// TIA Portal project "LabelProMax" (V16)

(* hardware
DEVICE "ET 200SP station_1"  ET 200SP-Station
   slot 0: "Rack_0"  Rack  6ES5 710-8MAx1
   slot 1: "PLC_label"  CPU 1512SP F-1 PN  6ES7 512-1SK01-0AB0  V2.8
      slot 32768: "PROFINET interface_1"  X1
         slot 32771: "Port_3"  X1 P3
   slot 2: "DI 8x24VDC HF_1"  DI 8x24VDC HF  6ES7 131-6BF00-0CA0  V1.2
      slot 1: "DI 8x24VDC HF_1"  DI 8x24VDC HF
   slot 3: "DI 8x24VDC HF_2"  DI 8x24VDC HF  6ES7 131-6BF00-0CA0  V1.2
      slot 1: "DI 8x24VDC HF_2"  DI 8x24VDC HF
   slot 4: "DQ 8x24VDC/0.5A HF_1"  DQ 8x24VDC/0.5A HF  6ES7 132-6BF00-0CA0  V1.2
      slot 1: "DQ 8x24VDC/0.5A HF_1"  DQ 8x24VDC/0.5A HF
   slot 5: "DQ 8x24VDC/0.5A HF_2"  DQ 8x24VDC/0.5A HF  6ES7 132-6BF00-0CA0  V1.2
      slot 1: "DQ 8x24VDC/0.5A HF_2"  DQ 8x24VDC/0.5A HF
   slot 6: "CM 4xIO-Link_1"  CM 4xIO-Link  6ES7 137-6BD00-0BA0  V2.1
      slot 1: "CM 4xIO-Link_1"  6ES7 137-6BD00-0BA0
   slot 7: "Server module_1"  Server module  6ES7 193-6PA00-0AA0  V1.0
      slot 1: "Server module_1"  Server module
   slot 127: "BA 2xRJ45"  BA 2xRJ45  6ES7 193-6AR00-0AA0  V0.0
      slot 32769: "Port_1"  X1 P1  6ES7 193-6AR00-0AA0
      slot 32770: "Port_2"  X1 P2  6ES7 193-6AR00-0AA0
DEVICE "HMI_label"  TP700 Comfort
   slot 0: "HMI_label"  TP700 Comfort  6AV2 124-0GC01-0AX0  16.0.0.0
   slot 1: "HMI_RT_1"  TP700 Comfort  6AV2 124-0GC01-0AX0  16.0.0.0
   slot 5: "HMI_label.IE_CP_1"  PROFINET Interface  16.0.0.0
      slot 1: "PROFINET Interface_1"  PROFINET Interface
         slot 1: "Port_1"  Port
         slot 2: "Port_2"  Port
   slot 7: "HMI_label.MPI/DP_CP_1"  MPI/DP Interface  16.0.0.0
*)

// ===== PLC "PLC_label"  CPU 1512SP F-1 PN =====

VAR_GLOBAL   // PLC tag table "Default tag table"
   "start" AT %I1.0 : Bool;   // 1=Start button pushed
   "stop" AT %I1.1 : Bool;   // 0=Stop button pushed (NC)
   "F1_F2" AT %I1.2 : Bool;   // 0=F1
   "reset" AT %I1.3 : Bool;   // 1=Reset button pushed
   "conv_centre" AT %I1.4 : Bool;   // 1=Carrier at conveyor centre
   "estop" AT %I1.5 : Bool;   // 0=Emergency stop button pushed (NC)
   "conv_start" AT %I1.6 : Bool;   // 1=Carrier at conveyor start
   "conv_end" AT %I1.7 : Bool;   // 1=Carrier at conveyor end
   "start_lamp" AT %Q1.0 : Bool;   // 1=Start lamp is lit
   "reset_lamp" AT %Q1.1 : Bool;   // 1=Reset lamp is lit
   "indicator_1" AT %Q1.2 : Bool;   // 1=Indicator Light 1 is lit
   "indicator_2" AT %Q1.3 : Bool;   // 1=Indicator Light 2 is lit
   "conv_fwd" AT %Q1.4 : Bool;   // 1=Move conveyor belt in clockwise rotation (to the right)
   "conv_bwd" AT %Q1.5 : Bool;   // 1=Move conveyor belt in counterclockwise rotation (to the left)
   "conv_inch" AT %Q1.6 : Bool;   // 1=Activate inch-travel of conveyor belt
   "stopper" AT %Q1.7 : Bool;   // 1=Move stopper cylinder to lower end position
END_VAR

VAR_GLOBAL   // PLC tag table "Tag table_1"
   "BG1" AT %I0.0 : Bool;
   "BG2" AT %I0.1 : Bool;
   "BG3" AT %I0.2 : Bool;
   "BG4" AT %I0.3 : Bool;
   "BG5" AT %I0.4 : Bool;
   "BG6" AT %I0.5 : Bool;
   "MB1" AT %Q0.0 : Bool;
   "MB3" AT %Q0.2 : Bool;
   "MB4" AT %Q0.3 : Bool;
   "MB5" AT %Q0.4 : Bool;
   "MB6" AT %Q0.5 : Bool;
   "MB7" AT %Q0.6 : Bool;
   "MA8" AT %Q0.7 : Bool;
END_VAR

DATA_BLOCK "base_Module_DB"   // DB1
{ S7_Optimized_Access := 'TRUE' }
VERSION : 0.1
// stored: InstanceOfName base_Module
"base_Module"
BEGIN
END_DATA_BLOCK

DATA_BLOCK "application_Module_DB"   // DB2
{ S7_Optimized_Access := 'TRUE' }
VERSION : 0.1
// stored: InstanceOfName application_Module
"application_Module"
BEGIN
END_DATA_BLOCK

DATA_BLOCK "Data_block_1"   // DB3
{ S7_Optimized_Access := 'TRUE' }
VERSION : 0.1
   VAR
      flag : Bool;
      state : Int;
      State1_Active : Bool;
      State2_Active : Bool;
      State3_Active : Bool;
      done : Bool;
      prev_done : Bool;
      "counter" : Int;
      run_timer : Real;
      prev_start : Bool;
      rfidDone : Bool;
      cycle_timer : TON_TIME;
      cycle_time_ms : DInt;
      total_runtime_ms : DInt;
      prev_rfidDone : Bool;
      timer_enable : Bool;
   END_VAR
BEGIN
END_DATA_BLOCK

DATA_BLOCK "LIOLink_RF200_ReadTag_DB"   // DB5
{ S7_Optimized_Access := 'FALSE' }
// stored: InstanceOfName LIOLink_RF200_ReadTag
"LIOLink_RF200_ReadTag"
BEGIN
END_DATA_BLOCK

DATA_BLOCK "RFID_Control"   // DB6
{ S7_Optimized_Access := 'TRUE' }
VERSION : 0.1
   VAR
      read : Bool := false;   // Execute a read of the RFID tag on rising edge
      write : Bool := false;
      length : Word := 16#1C;
      addrTag : Word := 16#00;
      hwID : Hw_SubModule := 261;
      portAddr : Int := 0;
      "version" : USInt := 11;
      readDone : Bool := false;
      writeDone : Bool := false;
      readPresence : Bool;
      writePresence : Bool;
   END_VAR
BEGIN
END_DATA_BLOCK

DATA_BLOCK "LIOLink_RF200_WriteTag_DB"   // DB7
{ S7_Optimized_Access := 'FALSE' }
// stored: InstanceOfName LIOLink_RF200_WriteTag
"LIOLink_RF200_WriteTag"
BEGIN
END_DATA_BLOCK

DATA_BLOCK "identData"   // DB8
{ S7_Optimized_Access := 'TRUE' }
VERSION : 0.1
   VAR
      readData : Array[0..31] of Byte;
      writeData : Array[0..31] of Byte;
   END_VAR
BEGIN
END_DATA_BLOCK

DATA_BLOCK "DB_MES_Comms"   // DB9
{ S7_Optimized_Access := 'TRUE' }
VERSION : 0.1
   VAR
      var1 : Bool;
      var2 : Int;
      var3 : Array[0..7] of Real;
      current_order_id : Int;
      station_state : Int;
      run_time : Real;
      total_count : Int;
      good_count : Int;
      completion_status : Bool;
      label_request : Bool;
      label_text : String[80];
      print_status : Bool;
      last_cycle_time : Real;
      cycle_done : Bool;
   END_VAR
BEGIN
END_DATA_BLOCK

DATA_BLOCK "state_Transition_Module_DB"   // DB10
{ S7_Optimized_Access := 'TRUE' }
VERSION : 0.1
// stored: InstanceOfName state_Transition_Module
"state_Transition_Module"
BEGIN
END_DATA_BLOCK

DATA_BLOCK "rfid_Current_Order_Module_DB"   // DB11
{ S7_Optimized_Access := 'TRUE' }
VERSION : 0.1
// stored: InstanceOfName rfid_Current_Order_Module
"rfid_Current_Order_Module"
BEGIN
END_DATA_BLOCK

FUNCTION_BLOCK "base_Module"   // FB1, GRAPH_PLUS
{ S7_Optimized_Access := 'TRUE' }
VERSION : 0.1
   VAR_INPUT
      OFF_SQ : Bool := false;   // Turn sequence off
      INIT_SQ : Bool := false;   // Set sequence to initial state
      ACK_EF : Bool := false;   // Acknowledge all errors and faults
      S_PREV : Bool := false;   // Output previous step in parameter S_NO
      S_NEXT : Bool := false;   // Indicate next step in parameter S_NO
      SW_AUTO : Bool := false;   // Automatic mode
      SW_TAP : Bool := false;   // Semiautomatic/switch with transition
      SW_TOP : Bool := false;   // Semiautomatic/ignore transition
      SW_MAN : Bool := false;   // Manual mode
      S_SEL : Int := 0;   // Select step to be output to S_NO
      S_ON : Bool := false;   // Activate step indicated in S_NO
      S_OFF : Bool := false;   // Deactivate step indicated S_NO
      T_PUSH : Bool := false;   // Enable transition to switch in semi automatic mode
   END_VAR
   VAR_OUTPUT
      S_NO : Int := 0;   // Step number
      S_MORE : Bool := false;   // More steps are available and can be shown in S_NO
      S_ACTIVE : Bool := false;   // Step indicated in S_NO is active
      ERR_FLT : Bool := false;   // Interlock or supervision group error
      AUTO_ON : Bool := false;   // Automatic mode is active
      TAP_ON : Bool := false;   // Semiautomatic mode/step with transition enabled
      TOP_ON : Bool := false;   // Semiautomatic mode/ignore transition enabled
      MAN_ON : Bool := false;   // Manual mode is active
   END_VAR
   VAR
      HMI_INFO : Array[0..8] of UInt;
      IF_PAR : G7_IfParPlus_V6;
      RT_DATA : G7_RTDataPlus_V6;   // Internal data area
      Trans1 : G7_TransitionPlus_V6;   // Transition structure
      Trans2 : G7_TransitionPlus_V6;   // Transition structure
      Trans3 : G7_TransitionPlus_V6;   // Transition structure
      Trans4 : G7_TransitionPlus_V6;   // Transition structure
      Trans5 : G7_TransitionPlus_V6;   // Transition structure
      Trans6 : G7_TransitionPlus_V6;   // Transition structure
      Trans7 : G7_TransitionPlus_V6;   // Transition structure
      Trans8 : G7_TransitionPlus_V6;   // Transition structure
      Trans9 : G7_TransitionPlus_V6;   // Transition structure
      Step1 : G7_StepPlus_V6;   // Step structure
      Step2 : G7_StepPlus_V6;   // Step structure
      Step3 : G7_StepPlus_V6;   // Step structure
      Step4 : G7_StepPlus_V6;   // Step structure
      Step5 : G7_StepPlus_V6;   // Step structure
      Step6 : G7_StepPlus_V6;   // Step structure
      Step7 : G7_StepPlus_V6;   // Step structure
      Step8 : G7_StepPlus_V6;   // Step structure
      Step9 : G7_StepPlus_V6;   // Step structure
      SINI : Array[0..1] of USInt;
      LSTT : Array[0..8] of USInt;
      ATAJ : Array[0..8] of USInt;
      ATAB : Array[0..8] of USInt;
      PSTT : Array[0..8] of USInt;
      NSTT : Array[0..8] of USInt;
      ASSJ : Array[0..8] of USInt;
      ASSB : Array[0..8] of USInt;
      PTTS : Array[0..8] of USInt;
      NTTS : Array[0..8] of USInt;
      SW_SQTS : Array[0..8] of USInt;
      SWITCH : Array[0..0] of USInt;
      TVX : Array[0..1] of USInt;
      TTX : Array[0..1] of USInt;
      TSX : Array[0..1] of USInt;
      S00X : Array[0..1] of USInt;
      SOFFX : Array[0..1] of USInt;
      SONX : Array[0..1] of USInt;
      SAX : Array[0..1] of USInt;
      SERRX : Array[0..9] of USInt;
      SMX : Array[0..9] of USInt;
      S0X : Array[0..9] of USInt;
      S1X : Array[0..9] of USInt;
      IL_ALARM_INST : Diag_Alarm;
      SUP_ALARM_INST : Diag_Alarm;
      STEP_TIME_ALARM_INST : Diag_Alarm;
      IEC_TIMER_INST : IEC_TIMER;
      TRANSACTION_FLAG : Bool := false;
   END_VAR
   // SINI[0] := 2;
   // LSTT[0] := 255;
   // LSTT[1] := 255;
   // LSTT[2] := 255;
   // ATAJ[1] := 1;
   // ATAJ[2] := 2;
   // ATAJ[3] := 3;
   // ATAB[1] := 1;
   // ATAB[2] := 2;
   // ATAB[3] := 3;
   // PSTT[1] := 1;
   // PSTT[2] := 2;
   // PSTT[3] := 5;
   // NSTT[0] := 1;
   // NSTT[1] := 6;
   // NSTT[2] := 3;
   // ASSJ[1] := 1;
   // ASSJ[2] := 2;
   // ASSJ[3] := 3;
   // ASSB[1] := 1;
   // ASSB[2] := 2;
   // ASSB[3] := 3;
   // PTTS[0] := 255;
   // PTTS[2] := 8;
   // PTTS[3] := 2;
   // NTTS[1] := 1;
   // NTTS[2] := 2;
   // NTTS[3] := 5;
   // TVX[0] := 16#1;
   // TTX[0] := 16#1;
   // TSX[0] := 16#1;
   // S00X[0] := 16#1;
   // SOFFX[0] := 16#1;
   // SONX[0] := 16#1;
   // SAX[0] := 16#1;
   // SERRX[0] := 16#1;
   // SMX[0] := 16#1;
   // S0X[0] := 16#1;
   // S1X[0] := 16#1;
   // LSTT[3] := 255;
   // ATAJ[4] := 4;
   // ATAB[4] := 4;
   // PSTT[4] := 4;
   // NSTT[3] := 4;
   // ASSJ[4] := 4;
   // ASSB[4] := 4;
   // PTTS[4] := 3;
   // NTTS[4] := 4;
   // LSTT[5] := 255;
   // ATAJ[5] := 5;
   // ATAB[5] := 5;
   // PSTT[5] := 3;
   // NSTT[5] := 5;
   // ASSJ[5] := 5;
   // ASSB[5] := 5;
   // PTTS[5] := 5;
   // NTTS[5] := 3;
   // LSTT[6] := 255;
   // ATAJ[6] := 6;
   // ATAB[6] := 6;
   // PSTT[6] := 6;
   // NSTT[6] := 7;
   // ASSJ[6] := 6;
   // ASSB[6] := 6;
   // PTTS[6] := 1;
   // NTTS[6] := 6;
   // LSTT[7] := 255;
   // LSTT[8] := 255;
   // ATAJ[7] := 7;
   // ATAJ[8] := 8;
   // ATAB[7] := 7;
   // ATAB[8] := 8;
   // PSTT[7] := 7;
   // PSTT[8] := 8;
   // NSTT[7] := 8;
   // NSTT[8] := 2;
   // ASSJ[7] := 7;
   // ASSJ[8] := 8;
   // ASSB[7] := 7;
   // ASSB[8] := 8;
   // PTTS[7] := 6;
   // PTTS[8] := 7;
   // NTTS[7] := 7;
   // NTTS[8] := 8;
BEGIN
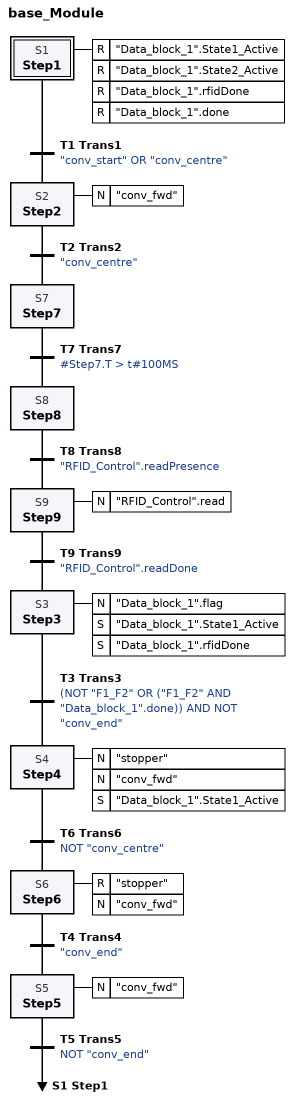
   // sequencer 1
   INITIAL_STEP Step1:   // S1, max time T#10S, warning time T#7S
              R    "Data_block_1".State1_Active
              R    "Data_block_1".State2_Active
              R    "Data_block_1".rfidDone
              R    "Data_block_1".done
   END_STEP
   TRANSITION Trans1 FROM Step1 TO Step2   // T1
      := "conv_start" OR "conv_centre";
   END_TRANSITION
   STEP Step2:   // S2, max time T#10S, warning time T#7S
              N    "conv_fwd"
   END_STEP
   TRANSITION Trans2 FROM Step2 TO Step7   // T2
      := "conv_centre";
   END_TRANSITION
   STEP Step3:   // S3, max time T#10S, warning time T#7S
              N    "Data_block_1".flag
              S    "Data_block_1".State1_Active
              S    "Data_block_1".rfidDone
   END_STEP
   TRANSITION Trans3 FROM Step3 TO Step4   // T3
      := (NOT "F1_F2" OR ("F1_F2" AND "Data_block_1".done)) AND NOT "conv_end";
   END_TRANSITION
   STEP Step4:   // S4, max time T#10S, warning time T#7S
              N    "stopper"
              N    "conv_fwd"
              S    "Data_block_1".State1_Active
   END_STEP
   TRANSITION Trans6 FROM Step4 TO Step6   // T6
      := NOT "conv_centre";
   END_TRANSITION
   STEP Step5:   // S5, max time T#10S, warning time T#7S
              N    "conv_fwd"
   END_STEP
   TRANSITION Trans5 FROM Step5 TO Step1   // T5, jump
      := NOT "conv_end";
   END_TRANSITION
   STEP Step6:   // S6, max time T#10S, warning time T#7S
              R    "stopper"
              N    "conv_fwd"
   END_STEP
   TRANSITION Trans4 FROM Step6 TO Step5   // T4
      := "conv_end";
   END_TRANSITION
   STEP Step7:   // S7, max time T#10S, warning time T#7S
   END_STEP
   TRANSITION Trans7 FROM Step7 TO Step8   // T7
      := #Step7.T > t#100MS;
   END_TRANSITION
   STEP Step8:   // S8, max time T#10S, warning time T#7S
   END_STEP
   TRANSITION Trans8 FROM Step8 TO Step9   // T8
      := "RFID_Control".readPresence;
   END_TRANSITION
   STEP Step9:   // S9, max time T#10S, warning time T#7S
              N    "RFID_Control".read
   END_STEP
   TRANSITION Trans9 FROM Step9 TO Step3   // T9
      := "RFID_Control".readDone;
   END_TRANSITION
END_FUNCTION_BLOCK

FUNCTION_BLOCK "application_Module"   // FB2, GRAPH_PLUS
{ S7_Optimized_Access := 'TRUE' }
VERSION : 0.1
   VAR_INPUT
      OFF_SQ : Bool := false;   // Turn sequence off
      INIT_SQ : Bool := false;   // Set sequence to initial state
      ACK_EF : Bool := false;   // Acknowledge all errors and faults
      S_PREV : Bool := false;   // Output previous step in parameter S_NO
      S_NEXT : Bool := false;   // Indicate next step in parameter S_NO
      SW_AUTO : Bool := false;   // Automatic mode
      SW_TAP : Bool := false;   // Semiautomatic/switch with transition
      SW_TOP : Bool := false;   // Semiautomatic/ignore transition
      SW_MAN : Bool := false;   // Manual mode
      S_SEL : Int := 0;   // Select step to be output to S_NO
      S_ON : Bool := false;   // Activate step indicated in S_NO
      S_OFF : Bool := false;   // Deactivate step indicated S_NO
      T_PUSH : Bool := false;   // Enable transition to switch in semi automatic mode
   END_VAR
   VAR_OUTPUT
      S_NO : Int := 0;   // Step number
      S_MORE : Bool := false;   // More steps are available and can be shown in S_NO
      S_ACTIVE : Bool := false;   // Step indicated in S_NO is active
      ERR_FLT : Bool := false;   // Interlock or supervision group error
      AUTO_ON : Bool := false;   // Automatic mode is active
      TAP_ON : Bool := false;   // Semiautomatic mode/step with transition enabled
      TOP_ON : Bool := false;   // Semiautomatic mode/ignore transition enabled
      MAN_ON : Bool := false;   // Manual mode is active
   END_VAR
   VAR
      HMI_INFO : Array[0..8] of UInt;
      IF_PAR : G7_IfParPlus_V6;
      RT_DATA : G7_RTDataPlus_V6;   // Internal data area
      Trans1 : G7_TransitionPlus_V6;   // Transition structure
      Trans2 : G7_TransitionPlus_V6;   // Transition structure
      Trans3 : G7_TransitionPlus_V6;   // Transition structure
      Trans4 : G7_TransitionPlus_V6;   // Transition structure
      Trans5 : G7_TransitionPlus_V6;   // Transition structure
      Trans6 : G7_TransitionPlus_V6;   // Transition structure
      Trans7 : G7_TransitionPlus_V6;   // Transition structure
      Trans8 : G7_TransitionPlus_V6;   // Transition structure
      Trans9 : G7_TransitionPlus_V6;   // Transition structure
      Trans10 : G7_TransitionPlus_V6;   // Transition structure
      Trans11 : G7_TransitionPlus_V6;   // Transition structure
      Step1 : G7_StepPlus_V6;   // Step structure
      Step2 : G7_StepPlus_V6;   // Step structure
      Step3 : G7_StepPlus_V6;   // Step structure
      Step4 : G7_StepPlus_V6;   // Step structure
      Step5 : G7_StepPlus_V6;   // Step structure
      Step6 : G7_StepPlus_V6;   // Step structure
      Step7 : G7_StepPlus_V6;   // Step structure
      Step8 : G7_StepPlus_V6;   // Step structure
      Step9 : G7_StepPlus_V6;   // Step structure
      Step10 : G7_StepPlus_V6;   // Step structure
      Step11 : G7_StepPlus_V6;   // Step structure
      SINI : Array[0..1] of USInt;
      LSTT : Array[0..10] of USInt;
      ATAJ : Array[0..10] of USInt;
      ATAB : Array[0..10] of USInt;
      PSTT : Array[0..10] of USInt;
      NSTT : Array[0..10] of USInt;
      ASSJ : Array[0..10] of USInt;
      ASSB : Array[0..10] of USInt;
      PTTS : Array[0..10] of USInt;
      NTTS : Array[0..10] of USInt;
      SW_SQTS : Array[0..10] of USInt;
      SWITCH : Array[0..0] of USInt;
      TVX : Array[0..1] of USInt;
      TTX : Array[0..1] of USInt;
      TSX : Array[0..1] of USInt;
      S00X : Array[0..1] of USInt;
      SOFFX : Array[0..1] of USInt;
      SONX : Array[0..1] of USInt;
      SAX : Array[0..1] of USInt;
      SERRX : Array[0..11] of USInt;
      SMX : Array[0..11] of USInt;
      S0X : Array[0..11] of USInt;
      S1X : Array[0..11] of USInt;
      IL_ALARM_INST : Diag_Alarm;
      SUP_ALARM_INST : Diag_Alarm;
      STEP_TIME_ALARM_INST : Diag_Alarm;
      IEC_TIMER_INST : IEC_TIMER;
      TRANSACTION_FLAG : Bool := false;
   END_VAR
   // SINI[0] := 2;
   // LSTT[0] := 255;
   // LSTT[1] := 255;
   // LSTT[2] := 255;
   // LSTT[3] := 255;
   // LSTT[4] := 255;
   // LSTT[5] := 255;
   // LSTT[6] := 255;
   // LSTT[7] := 255;
   // LSTT[8] := 255;
   // LSTT[9] := 255;
   // ATAJ[1] := 1;
   // ATAJ[2] := 2;
   // ATAJ[3] := 3;
   // ATAJ[4] := 4;
   // ATAJ[5] := 5;
   // ATAJ[6] := 6;
   // ATAJ[7] := 7;
   // ATAJ[8] := 8;
   // ATAJ[9] := 9;
   // ATAJ[10] := 10;
   // ATAB[1] := 1;
   // ATAB[2] := 2;
   // ATAB[3] := 3;
   // ATAB[4] := 4;
   // ATAB[5] := 5;
   // ATAB[6] := 6;
   // ATAB[7] := 7;
   // ATAB[8] := 8;
   // ATAB[9] := 9;
   // ATAB[10] := 10;
   // PSTT[1] := 1;
   // PSTT[2] := 2;
   // PSTT[3] := 3;
   // PSTT[4] := 4;
   // PSTT[5] := 5;
   // PSTT[6] := 6;
   // PSTT[7] := 7;
   // PSTT[8] := 8;
   // PSTT[9] := 9;
   // PSTT[10] := 10;
   // NSTT[0] := 1;
   // NSTT[1] := 2;
   // NSTT[2] := 3;
   // NSTT[3] := 4;
   // NSTT[4] := 5;
   // NSTT[5] := 6;
   // NSTT[6] := 7;
   // NSTT[7] := 8;
   // NSTT[8] := 9;
   // NSTT[9] := 10;
   // ASSJ[1] := 1;
   // ASSJ[2] := 2;
   // ASSJ[3] := 3;
   // ASSJ[4] := 4;
   // ASSJ[5] := 5;
   // ASSJ[6] := 6;
   // ASSJ[7] := 7;
   // ASSJ[8] := 8;
   // ASSJ[9] := 9;
   // ASSJ[10] := 10;
   // ASSB[1] := 1;
   // ASSB[2] := 2;
   // ASSB[3] := 3;
   // ASSB[4] := 4;
   // ASSB[5] := 5;
   // ASSB[6] := 6;
   // ASSB[7] := 7;
   // ASSB[8] := 8;
   // ASSB[9] := 9;
   // ASSB[10] := 10;
   // PTTS[0] := 255;
   // PTTS[2] := 1;
   // PTTS[3] := 2;
   // PTTS[4] := 3;
   // PTTS[5] := 4;
   // PTTS[6] := 5;
   // PTTS[7] := 6;
   // PTTS[8] := 7;
   // PTTS[9] := 8;
   // PTTS[10] := 9;
   // NTTS[1] := 1;
   // NTTS[2] := 2;
   // NTTS[3] := 3;
   // NTTS[4] := 4;
   // NTTS[5] := 5;
   // NTTS[6] := 6;
   // NTTS[7] := 7;
   // NTTS[8] := 8;
   // NTTS[9] := 9;
   // NTTS[10] := 10;
   // TVX[0] := 16#1;
   // TTX[0] := 16#1;
   // TSX[0] := 16#1;
   // S00X[0] := 16#1;
   // SOFFX[0] := 16#1;
   // SONX[0] := 16#1;
   // SAX[0] := 16#1;
   // SERRX[0] := 16#1;
   // SMX[0] := 16#1;
   // S0X[0] := 16#1;
   // S1X[0] := 16#1;
BEGIN
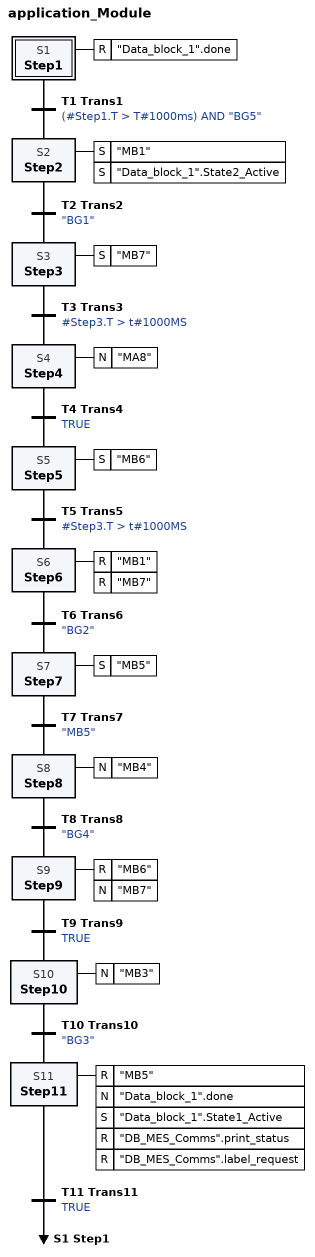
   // sequencer 1
   INITIAL_STEP Step1:   // S1, max time T#10S, warning time T#7S
              R    "Data_block_1".done
   END_STEP
   TRANSITION Trans1 FROM Step1 TO Step2   // T1
      := (#Step1.T > T#1000ms) AND "BG5";
   END_TRANSITION
   STEP Step2:   // S2, max time T#10S, warning time T#7S
              S    "MB1"
              S    "Data_block_1".State2_Active
   END_STEP
   TRANSITION Trans2 FROM Step2 TO Step3   // T2
      := "BG1";
   END_TRANSITION
   STEP Step3:   // S3, max time T#10S, warning time T#7S
              S    "MB7"
   END_STEP
   TRANSITION Trans3 FROM Step3 TO Step4   // T3
      := #Step3.T > t#1000MS;
   END_TRANSITION
   STEP Step4:   // S4, max time T#10S, warning time T#7S
              N    "MA8"
   END_STEP
   TRANSITION Trans4 FROM Step4 TO Step5   // T4
      := TRUE;
   END_TRANSITION
   STEP Step5:   // S5, max time T#10S, warning time T#7S
              S    "MB6"
   END_STEP
   TRANSITION Trans5 FROM Step5 TO Step6   // T5
      := #Step3.T > t#1000MS;
   END_TRANSITION
   STEP Step6:   // S6, max time T#10S, warning time T#7S
              R    "MB1"
              R    "MB7"
   END_STEP
   TRANSITION Trans6 FROM Step6 TO Step7   // T6
      := "BG2";
   END_TRANSITION
   STEP Step7:   // S7, max time T#10S, warning time T#7S
              S    "MB5"
   END_STEP
   TRANSITION Trans7 FROM Step7 TO Step8   // T7
      := "MB5";
   END_TRANSITION
   STEP Step8:   // S8, max time T#10S, warning time T#7S
              N    "MB4"
   END_STEP
   TRANSITION Trans8 FROM Step8 TO Step9   // T8
      := "BG4";
   END_TRANSITION
   STEP Step9:   // S9, max time T#10S, warning time T#7S
              R    "MB6"
              N    "MB7"
   END_STEP
   TRANSITION Trans9 FROM Step9 TO Step10   // T9
      := TRUE;
   END_TRANSITION
   STEP Step10:   // S10, max time T#10S, warning time T#7S
              N    "MB3"
   END_STEP
   TRANSITION Trans10 FROM Step10 TO Step11   // T10
      := "BG3";
   END_TRANSITION
   STEP Step11:   // S11, max time T#10S, warning time T#7S
              R    "MB5"
              N    "Data_block_1".done
              S    "Data_block_1".State1_Active
              R    "DB_MES_Comms".print_status
              R    "DB_MES_Comms".label_request
   END_STEP
   TRANSITION Trans11 FROM Step11 TO Step1   // T11, jump
      := TRUE;
   END_TRANSITION
END_FUNCTION_BLOCK

FUNCTION_BLOCK "state_Transition_Module"   // FB4, SCL
{ S7_Optimized_Access := 'TRUE' }
VERSION : 0.1
BEGIN
   IF "Data_block_1".State2_Active THEN
       "Data_block_1".state := 2;
       "DB_MES_Comms".station_state := "Data_block_1".state;
   ELSIF "Data_block_1".State1_Active THEN
       "Data_block_1".state := 1;
       "DB_MES_Comms".station_state := "Data_block_1".state;
   ELSE
       "Data_block_1".state := 0;
       "DB_MES_Comms".station_state := "Data_block_1".state;
   END_IF;
END_FUNCTION_BLOCK

ORGANIZATION_BLOCK "Main"   // OB1, LAD, ProgramCycle
TITLE = "Main Program Sweep (Cycle)"
{ S7_Optimized_Access := 'TRUE' }
VERSION : 0.1
   VAR_INPUT
      Initial_Call : Bool;   // Initial call of this OB
      Remanence : Bool;   // =True, if remanent data are available
   END_VAR
   VAR_TEMP
      run_time_ms : Real;
   END_VAR
BEGIN

REGION Network 1: Execution of Converyor belt start stop logic in Block_1 [FB1]
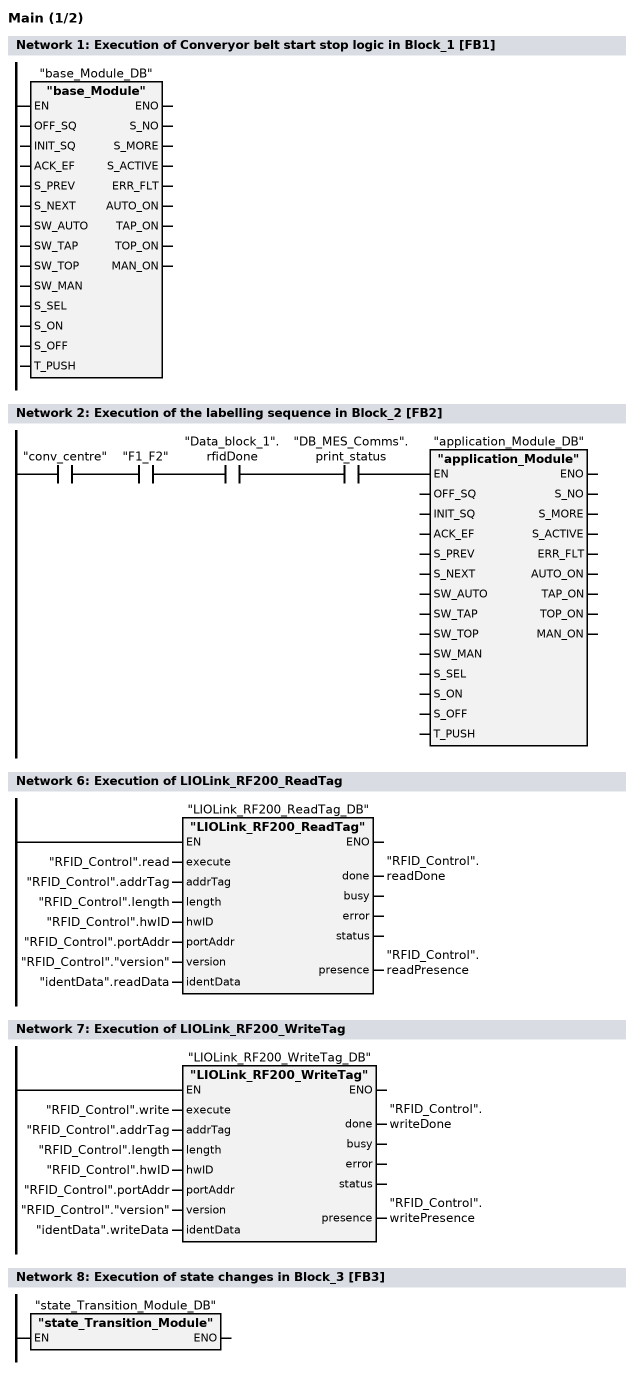
   RUNG wire#powerrail
      "base_Module_DB"(OFF_SQ :=, INIT_SQ :=, ACK_EF :=, S_PREV :=, S_NEXT :=, SW_AUTO :=, SW_TAP :=, SW_TOP :=, SW_MAN :=, S_SEL :=, S_ON :=, S_OFF :=, T_PUSH :=, S_NO =>, S_MORE =>, S_ACTIVE =>, ERR_FLT =>, AUTO_ON =>, TAP_ON =>, TOP_ON =>, MAN_ON =>)
   END_RUNG
   // the same network as SCL:
   "base_Module_DB"();   // "base_Module"
END_REGION

REGION Network 2: Execution of the labelling sequence in Block_2 [FB2]
   RUNG wire#powerrail
      Contact( "conv_centre" )
      Contact( "F1_F2" )
      Contact( "Data_block_1".rfidDone )
      Contact( "DB_MES_Comms".print_status )
      "application_Module_DB"(OFF_SQ :=, INIT_SQ :=, ACK_EF :=, S_PREV :=, S_NEXT :=, SW_AUTO :=, SW_TAP :=, SW_TOP :=, SW_MAN :=, S_SEL :=, S_ON :=, S_OFF :=, T_PUSH :=, S_NO =>, S_MORE =>, S_ACTIVE =>, ERR_FLT =>, AUTO_ON =>, TAP_ON =>, TOP_ON =>, MAN_ON =>)
   END_RUNG
   // the same network as SCL:
   IF "conv_centre" AND "F1_F2" AND "Data_block_1".rfidDone AND "DB_MES_Comms".print_status THEN
       "application_Module_DB"();   // "application_Module"
   END_IF;
END_REGION

REGION Network 3 (SCL): Total Count
   IF "Data_block_1".State1_Active AND NOT "Data_block_1".prev_start AND "F1_F2" = TRUE THEN

       "DB_MES_Comms".total_count := "DB_MES_Comms".total_count + 1;

   END_IF;

   "Data_block_1".prev_start := "Data_block_1".State1_Active;
END_REGION

REGION Network 4 (SCL): Good Count
   IF "Data_block_1".done AND NOT "Data_block_1".prev_done AND "F1_F2" = TRUE THEN

       "DB_MES_Comms".good_count := "DB_MES_Comms".good_count + 1;

   END_IF;

   "Data_block_1".prev_done := "Data_block_1".done;
END_REGION

REGION Network 5 (SCL): Completion Status of the orders sent by MES (not in reality\)
   IF "DB_MES_Comms".total_count >= 10 THEN
       "DB_MES_Comms".completion_status := TRUE;
   ELSE
       "DB_MES_Comms".completion_status := FALSE;
   END_IF;
END_REGION

REGION Network 6: Execution of LIOLink_RF200_ReadTag
   RUNG wire#powerrail
      "LIOLink_RF200_ReadTag_DB"(execute := "RFID_Control".read, addrTag := "RFID_Control".addrTag, length := "RFID_Control".length, hwID := "RFID_Control".hwID, portAddr := "RFID_Control".portAddr, "version" := "RFID_Control"."version", identData := "identData".readData, done => "RFID_Control".readDone, busy =>, error =>, status =>, presence => "RFID_Control".readPresence)
   END_RUNG
   // the same network as SCL:
   "LIOLink_RF200_ReadTag_DB"(execute := "RFID_Control".read,   // "LIOLink_RF200_ReadTag"
                           addrTag := "RFID_Control".addrTag,
                           length := "RFID_Control".length,
                           hwID := "RFID_Control".hwID,
                           portAddr := "RFID_Control".portAddr,
                           "version" := "RFID_Control"."version",
                           identData := "identData".readData,
                           done => "RFID_Control".readDone,
                           presence => "RFID_Control".readPresence);
END_REGION

REGION Network 7: Execution of LIOLink_RF200_WriteTag
   RUNG wire#powerrail
      "LIOLink_RF200_WriteTag_DB"(execute := "RFID_Control".write, addrTag := "RFID_Control".addrTag, length := "RFID_Control".length, hwID := "RFID_Control".hwID, portAddr := "RFID_Control".portAddr, "version" := "RFID_Control"."version", identData := "identData".writeData, done => "RFID_Control".writeDone, busy =>, error =>, status =>, presence => "RFID_Control".writePresence)
   END_RUNG
   // the same network as SCL:
   "LIOLink_RF200_WriteTag_DB"(execute := "RFID_Control".write,   // "LIOLink_RF200_WriteTag"
                           addrTag := "RFID_Control".addrTag,
                           length := "RFID_Control".length,
                           hwID := "RFID_Control".hwID,
                           portAddr := "RFID_Control".portAddr,
                           "version" := "RFID_Control"."version",
                           identData := "identData".writeData,
                           done => "RFID_Control".writeDone,
                           presence => "RFID_Control".writePresence);
END_REGION

REGION Network 8: Execution of state changes in Block_3 [FB3]
   RUNG wire#powerrail
      "state_Transition_Module_DB"()
   END_RUNG
   // the same network as SCL:
   "state_Transition_Module_DB"();   // "state_Transition_Module"
END_REGION

REGION Network 9 (SCL): Start Timer on RFID Done
   IF "Data_block_1".rfidDone AND NOT "Data_block_1".prev_rfidDone THEN
       "Data_block_1".timer_enable := TRUE;
   END_IF;

   "Data_block_1".prev_rfidDone := "Data_block_1".rfidDone;
END_REGION

REGION Network 10 (SCL): Cycle Timer (Controlled)
   "Data_block_1".cycle_timer(
                              IN := "Data_block_1".timer_enable,
                              PT := T#9999s
   );
END_REGION

REGION Network 11 (SCL): Stop Timer + Accumulate Runtime
   IF "Data_block_1".done AND NOT "Data_block_1".prev_done THEN

       "Data_block_1".timer_enable := false;

       "Data_block_1".cycle_time_ms := "Data_block_1".cycle_timer.ET;

       "Data_block_1".total_runtime_ms := "Data_block_1".total_runtime_ms + "Data_block_1".cycle_time_ms;

       "DB_MES_Comms".last_cycle_time := DINT_TO_REAL("Data_block_1".cycle_time_ms) / 1000.0;

       "DB_MES_Comms".cycle_done := TRUE;

   END_IF;

   "Data_block_1".prev_done := "Data_block_1".done;
END_REGION

REGION Network 12 (SCL): Reset cycle_done Signal
   IF "DB_MES_Comms".cycle_done THEN
       "DB_MES_Comms".cycle_done := FALSE;
   END_IF;
END_REGION

REGION Network 13 (SCL): MES Publish
   "DB_MES_Comms".run_time := DINT_TO_REAL("Data_block_1".total_runtime_ms) / 1000.0;
   "DB_MES_Comms".station_state := "Data_block_1".state;
END_REGION

REGION Network 14: Activate DB_MES_Comms.label_request when LIO...ReadTag_DB.done is true and DB...ms.print_status is false
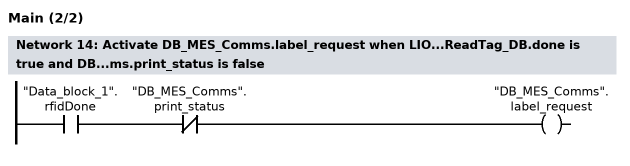
   RUNG wire#powerrail
      Contact( "Data_block_1".rfidDone )
      I_Contact( "DB_MES_Comms".print_status )
      Coil( "DB_MES_Comms".label_request )
   END_RUNG
   // the same network as SCL:
   "DB_MES_Comms".label_request := "Data_block_1".rfidDone AND NOT "DB_MES_Comms".print_status;
END_REGION
END_ORGANIZATION_BLOCK

// folder: LIOLink/S7-1200/1500/Device-specific blocks/SIMATIC RF200

FUNCTION_BLOCK "LIOLink_RF200_ReadTag"   // FB3, SCL
TITLE = LIOLink_RF200_ReadTag
{ S7_Optimized_Access := 'FALSE' }
// Reads tags from SIMATIC RF200 readers via IO-Link
   VAR_INPUT
      execute : Bool;   // Execute function
      addrTag : Word;   // Start address of data on tag
      length : Word;   // Length of data to be read
      hwID : Hw_SubModule;   // Hardware identifier of IO-Link communication module
      portAddr : Int;   // Start address of port
      "version" : USInt := 11;   // IO-Link version of the reader; 11: IO-Link V1.1, 10: IO-Link V1.0
   END_VAR
   VAR_OUTPUT
      done : Bool;
      busy : Bool;
      error : Bool;
      status : DWord;
      statusWord AT status : Array[0..1] of Word;
      presence : Bool;
   END_VAR
   VAR_IN_OUT
      identData : Variant;
   END_VAR
   VAR
      statPae : Array[0..27] of Byte;
      statStatusByte : Byte;
      statStatusBit AT statStatusByte : Array[0..7] of Bool;
      statPresence : Bool;
      statState : Int;
      statIdleState : Int;
      statTelegramState : Int := 1;
      statReadState : Int := 2;
      statErrorState : Int := 3;
      statAddr : Word;
      statAddrRead AT statAddr : Array[0..1] of Byte;
      statOffset : Int;
      statExecuteReq : Bool;
      statLength : DInt;
      statDat : Array[0..31] of Byte;
      statRecDat : Array[0..31] of Byte;
      statAddrOffset : Int;
      statPresenceFF : Bool;
      InstTonrTime : TONR_TIME;
      statTimerIn : Bool;
      statTimerR : Bool;
      statTimerPt : Time := t#5s;
      statReadData : Array[0..1999] of Byte;
      statCountCopyPae : DInt;
      statBusy : Bool;
      statDone : Bool;
      statReturnMoveBlkVar : Int;
      statDiffToIOsizeNetto : Int;
      InstSetIoPart : SETIO_PART;
      statIoPartError : Bool;
      statIoPartStatus : DWord;
      InstGetIoPart : GETIO_PART;
      statIOsize : USInt;
      statIOsizeNetto : USInt;
   END_VAR
   VAR_TEMP
      tempError : Bool;
      tempStatus : DWord;
      tempStatus_W AT tempStatus : Array[0..1] of Word;
   END_VAR
   VAR CONSTANT
      IOL_V10 : USInt := 10;   // Identifier IO-Link version 1.0
      IOL_V11 : USInt := 11;   // Identifier IO-Link version 1.1
      LEN_DATA_V10 : USInt := 8;   // Length of user data for IO-Link version 1.0
      LEN_DATA_V11 : USInt := 32;   // Length of user data for IO-Link version 1.1
   END_VAR
BEGIN
   REGION BLOCK INFO HEADER
     //===============================================================================
     // Siemens / (c)Copyright 2020
     //-------------------------------------------------------------------------------
     // Title:            LIOLink_RF200_ReadTag
     // Function:         Reads tags from SIMATIC RF200 readers via IO-Link
     // Library:          LIOLink
     // Author:           Siemens Industry Online Support
     // Tested with:      CPU 1513-1 PN FW 2.8
     // Engineering:      TIA Portal V16
     // Restrictions:     --
     // Requirements:     --
     //-------------------------------------------------------------------------------
     // Change log table:
     // Version  | Date       | Expert in charge       | Changes applied
     //----------|------------|------------------------|------------------------------
     // 01.00.00 | 01.07.2013 | Online Support         | First release
     // 01.01.00 | 01.12.2016 | Online Support         | Upgraded to TIA Portal V14
     // 02.00.00 | 01.09.2017 | Online Support         | Upgraded to TIA Portal V14 SP1
     //                                                | Implemented Programming styleguide
     //                                                | Added support for IO-Link V1.1 readers
     // 02.01.00 | 01.12.2017 | Online Support         | Bug fixes and performance improvements
     // 02.02.00 | 01.03.2020 | Online Support         | Upgraded to TIA Portal V16
     // 02.03.00 | 22.09.2020 | Online Support         | Integrated FB into LIOLink library
     //                                                | Renamed FB to LIOLink_RF200_ReadTag
     //                                                | Combined FBs for IO-Link V1.0 and V1.1
     //                                                | Minor bug fixes
     //===============================================================================
   END_REGION

   IF #version = #IOL_V11 THEN                               //determine IO-Link reader version (1.0/1.1) to set offsets
       #statIOsize := #LEN_DATA_V11;
       #statIOsizeNetto := #LEN_DATA_V11 - 4;
   ELSE
       #statIOsize := #LEN_DATA_V10;
       #statIOsizeNetto := #LEN_DATA_V10 - 4;
   END_IF;

   #statAddrOffset := #portAddr;                           //start adress of port
   #InstGetIoPart(ID     := #hwID,
                  OFFSET := #statAddrOffset,
                  LEN    := #statIOsize,
                  STATUS => #statIoPartStatus,
                  ERROR  => #statIoPartError,
                  INPUTS := #statRecDat);

   #statStatusByte := #statRecDat[0];         //Status Byte
   #statPresence := #statStatusBit[5];                     //Presence bit. Transponder on field
   #presence := #statPresence;

   IF NOT #execute THEN
       #statDone := false;
       #statBusy := false;
       #done := false;
       #busy := false;
       #error := false;
       #status := 0;
   ELSE
       #done := #statDone;
       #busy := #statBusy;
   END_IF;

   IF #execute AND #execute <> #statExecuteReq THEN        //Positive edge for d#reading of data
       IF NOT #statBusy THEN
           #statAddr := #addrTag;                                    //Transpoder Address
           #statDiffToIOsizeNetto := WORD_TO_INT(#length) MOD #statIOsizeNetto;
           #statLength := #length;                                 //Length of read Dat
           #statBusy := TRUE;
           #statDone := FALSE;                                     //reset all the output parameters                                   
           #error := FALSE;
           #status := 0;
           #statOffset := 0;                                       //offset of puffer must be reseted
           #statState := #statReadState;                           //next step >> send read command
           #statCountCopyPae := 0;
           FILL_BLK(IN    := 0,                                    //Reset read buffer
                    COUNT := CountOfElements(#identData),
                    OUT   => #statReadData[0]);
       ELSE
           #tempStatus_W[1] := 16#8102;                            //block is still active
           #tempStatus_W[0] := 16#0001;                            //Error identifier for block errors
           #status := #tempStatus;
           #statState := #statErrorState;
       END_IF;
       IF #length < 0 THEN
           #tempStatus_W[1] := 16#8104;                             //length too short
           #tempStatus_W[0] := 16#0001;                             //identifier rfid errors
           #status := #tempStatus;
           #statState := #statErrorState;
       END_IF;
   END_IF;
   #statExecuteReq := #execute;

   IF NOT #presence AND #presence <> #statPresenceFF THEN   //the tag has left the antenna  field
       IF NOT #statDone THEN
           #statTimerIn := true;                              //wait 5 sec
           #statTimerR := false;
       END_IF;
   END_IF;
   #statPresenceFF := #presence;
   IF #presence THEN
       #statTimerR := true;
       #statTimerIn := false;
   END_IF;
   //-----------------------------------------------------------------------------------------------------//
   //------------------------------------------start of state machine------------------------------------//
   //-----------------------------------------------------------------------------------------------------//
   CASE #statState OF
       0://IDLE
           #statBusy := false;
           #statTimerIn := false;

           (*
           // #statAdr := 0;
           // #statDat[0] := 16#0;                      //Set read command
           // #statDat[2] := #statAdrRead[0];             //Adr-H
           // #statDat[3] := #statAdrRead[1];             //Adr-L
           // #InstSetIoPart(ID:=#hwId,
           //                OFFSET:=#statAdrOffset,
           //                LEN:=8,
           //                STATUS=>#statIoPartStatus,
           //                ERROR=>#statIoPartError,
           //                OUTPUTS:=#statDat);
           *)
           //-------------------------------------------------Read state------------------------------------------//
           //---------------------------------------------sent read command---------------------------------------//
           //-----------------------------------------------------------------------------------------------------//

       2://Read_state

           IF #statLength > 0 THEN
               #statDat[0] := 16#2;                      //Set read command
               #statDat[2] := #statAddrRead[0];             //Adr-H
               #statDat[3] := #statAddrRead[1];             //Adr-L
           END_IF;

           IF NOT #statIoPartError THEN
               #statState := #statTelegramState;                           //Telegram: Edit the read data
           END_IF;


           //-----------------------------------------------Telegram state----------------------------------------//
           //---------------------------------------------edit received data--------------------------------------//
           //-----------------------------------------------------------------------------------------------------//  

       1://Telegram_state

           IF #statLength > 0 THEN                      //Only when length of data>0 can continue  
               IF #statStatusBit[6] THEN                                   //IF RFID error has occured
                   #tempStatus_W[1] := #statRecDat[1];    //error_RFID
                   #tempStatus_W[0] := 16#0011;                            //Error identifier for RFID errors
                   #status := #tempStatus;
                   #statState := #statErrorState;
               END_IF;

               //-------------------------- read command is ready------------------------------------------------//

               IF #statStatusBit[7] AND #statStatusBit[1] THEN
                   IF #statRecDat[2] = #statAddrRead[0]
                       AND #statRecDat[3] = #statAddrRead[1]
                   THEN //received ADR must be ==sent ADR
                       #statReturnMoveBlkVar := MOVE_BLK_VARIANT(SRC := #statRecDat,
                                                                 COUNT := #statIOsizeNetto,
                                                                 SRC_INDEX := 4,
                                                                 DEST_INDEX := 0,
                                                                 DEST => #statPae);

                       IF NOT #statIoPartError THEN
                           IF #statCountCopyPae = 0 THEN    //copy the #statIOsizeNet Bytes in 
                               IF #statLength >= #statIOsizeNetto THEN
                                   IF #statLength <> #length THEN
                                       #statAddr := INT_TO_WORD(WORD_TO_INT(#statAddr) + #statIOsizeNetto);
                                   END_IF;
                                   #statState := #statReadState;
                                   #statCountCopyPae := #statIOsizeNetto;
                               ELSE
                                   IF #statStatusBit[7] AND NOT #statStatusBit[6] THEN
                                       IF #statDiffToIOsizeNetto <> 0 THEN
                                           #statCountCopyPae := #statDiffToIOsizeNetto;
                                           #statAddr := INT_TO_WORD(WORD_TO_INT(#statAddr) + #statIOsizeNetto);
                                           #statState := #statReadState;
                                       ELSE
                                           #statCountCopyPae := #statIOsizeNetto;
                                       END_IF;
                                   ELSE
                                       #statState := #statIdleState;
                                   END_IF;
                               END_IF;
                           ELSE
                               #statReturnMoveBlkVar := MOVE_BLK_VARIANT(SRC := #statPae,
                                                                         COUNT := DINT_TO_UDINT(#statCountCopyPae),
                                                                         SRC_INDEX := 0,
                                                                         DEST_INDEX := #statOffset,
                                                                         DEST => #statReadData);
                               IF #statReturnMoveBlkVar = 0 THEN
                                   #statCountCopyPae := 0;
                                   #statOffset := #statOffset + #statIOsizeNetto;
                                   #statLength := #statLength - #statIOsizeNetto;
                               END_IF;
                           END_IF;
                       ELSE
                           #tempStatus_W[1] := DWORD_TO_WORD(#statIoPartStatus);                 //Error has to BLKMOV occured
                           #tempStatus_W[0] := 16#0001;                           //functions-Error identifier
                           #status := #tempStatus;
                           #statState := #statErrorState;
                       END_IF;
                   END_IF;
               END_IF;
               #InstSetIoPart(ID      := #hwID,
                              OFFSET  := #statAddrOffset,
                              LEN     := #statIOsize,
                              STATUS  => #statIoPartStatus,
                              ERROR   => #statIoPartError,
                              OUTPUTS := #statDat);

               IF #statIoPartError THEN
                   #tempStatus_W[1] := DWORD_TO_WORD(#statIoPartStatus);   //Error has to BLKMOV occured
                   #tempStatus_W[0] := 16#0001;                            //functions-Error identifier
                   #status := #tempStatus;
                   #statState := #statErrorState;
               END_IF;

           ELSE
               VariantPut(SRC := #statReadData,
                          DST := #identData);
               #statState := #statIdleState;
               #statBusy := false;
               #statDone := TRUE;

               //Reset read command
               #statDat[0] := 16#0;

               #InstSetIoPart(ID      := #hwID,
                              OFFSET  := #statAddrOffset,
                              LEN     := #statIOsize,
                              STATUS  => #statIoPartStatus,
                              ERROR   => #statIoPartError,
                              OUTPUTS := #statDat);
           END_IF;

           //------------------------------------------------------------------------------------------------------------//
           //-------------------------------------------------Error state------------------------------------------------//
           //---------------------------------------------error has occured----------------------------------------------//

       3://Error_State
           #tempError := TRUE;
           #statBusy := false;
           #error := #tempError;
           #statDone := false;
           #statTimerIn := false;
           #statTimerR := true;
           #statState := #statIdleState;
           #status := #tempStatus;

           //Reset read command
           #statDat[0] := 16#0;

           #InstSetIoPart(ID      := #hwID,
                          OFFSET  := #statAddrOffset,
                          LEN     := #statIOsize,
                          STATUS  => #statIoPartStatus,
                          ERROR   => #statIoPartError,
                          OUTPUTS := #statDat);
   END_CASE;

   //------------------------------------------------------------------------------------------------------------//
   //-------------------------------------------------Timer------------------------------------------------------//
   //------------------------------------------------------------------------------------------------------------//

   #InstTonrTime(IN := #statTimerIn,                  //this timer will start, if the tag has left the antenna field
                 R  := #statTimerR,
                 PT := #statTimerPt);
   IF #InstTonrTime.Q THEN                           //error has occured. No tag on field during the 5 sec.
       #tempStatus_W[1] := 16#8101;                           //tag has left the field
       #tempStatus_W[0] := 16#0001;                           //identifier rfid errors
       #status := #tempStatus;
       #statState := #statErrorState;
   END_IF;
END_FUNCTION_BLOCK

FUNCTION_BLOCK "LIOLink_RF200_WriteTag"   // FB5, SCL
TITLE = LIOLink_RF200_WriteTag
{ S7_Optimized_Access := 'FALSE' }
// Writes tags on SIMATIC RF200 readers via IO-Link
   VAR_INPUT
      execute : Bool;   // Execute function
      addrTag : Word;   // Start address of data on tag
      length : Word;   // Length of data to be written
      hwID : Hw_SubModule;   // Hardware identifier of IO-Link communication module
      portAddr : Int;   // Start address of port
      "version" : USInt := 11;   // IO-Link version of the reader; 11: IO-Link V1.1, 10: IO-Link V1.0
   END_VAR
   VAR_OUTPUT
      done : Bool;   // Ready
      busy : Bool;   // Block active
      error : Bool;   // Error has occured
      status : DWord;   // Error Status
      statusWord AT status : Array[0..1] of Word;
      presence : Bool;   // Tag on antenna field
   END_VAR
   VAR_IN_OUT
      identData : Variant;   // Data to write in
   END_VAR
   VAR
      instTonR : TONR_TIME;   // Timer 2
      statNState : Int;   // current state
      statTimerIn : Bool;   // Timer 2 parameters
      statTimerR : Bool;
      statTimerPt : Time := T#5s;
      statTelegramState : Int := 1;   // Edit state
      statWriteState : Int := 2;   // Write Command state
      statErrorState : Int := 3;   // Error state
      statIdleState : Int;   // first state
      statAddrOffset : Int;
      statStatusByte : Byte;   // first received Byte from process image
      statStatusBits AT statStatusByte : Array[0..7] of Bool;
      statDat : Array[0..31] of Byte;   // sent data
      statRecDat : Array[0..31] of Byte;   // writing data
      statPresenceBit : Bool;   // Presence bit
      statExecuteReq : Bool;
      statLength : DInt;
      statAddr : Word;   // address of Tag
      statAddrWrite AT statAddr : Array[0..1] of Byte;
      statWriteOffset : Int;
      statPresenceFf : Bool;
      statWriteData : Array[0..1999] of Byte;
      statAddrTag : Int;
      statDiffToIOsizeNetto : Int;
      statBytemove : Int;
      statDone : Bool;
      statBusy : Bool;
      InstSetIoPart : SETIO_PART;
      statIoPartError : Bool;
      statIoPartStatus : DWord;
      InstGetIoPart : GETIO_PART;
      statReturnMoveBlkVar : Int;
      statIOsize : USInt;
      statIOsizeNetto : USInt;
   END_VAR
   VAR_TEMP
      tempError : Bool;
      tempStatus : DWord;
      tempStatus_W AT tempStatus : Array[0..1] of Word;
   END_VAR
   VAR CONSTANT
      IOL_V10 : USInt := 10;   // Identifier IO-Link version 1.0
      IOL_V11 : USInt := 11;   // Identifier IO-Link version 1.1
      LEN_DATA_V10 : USInt := 8;   // Length of user data for IO-Link version 1.0
      LEN_DATA_V11 : USInt := 32;   // Length of user data for IO-Link version 1.1
   END_VAR
   // statRecDat[2] := 16#ff;
   // statRecDat[3] := 16#ff;
BEGIN
   REGION BLOCK INFO HEADER
     //===============================================================================
     // Siemens / (c)Copyright 2020
     //-------------------------------------------------------------------------------
     // Title:            LIOLink_RF200_WriteTag
     // Function:         Writes tags on SIMATIC RF200 readers via IO-Link
     // Library:          LIOLink
     // Author:           Siemens Industry Online Support
     // Tested with:      CPU 1513-1 PN FW 2.8
     // Engineering:      TIA Portal V16
     // Restrictions:     --
     // Requirements:     --
     //-------------------------------------------------------------------------------
     // Change log table:
     // Version  | Date       | Expert in charge       | Changes applied
     //----------|------------|------------------------|------------------------------
     // 01.00.00 | 01.03.2015 | Online Support         | First release
     // 01.01.00 | 01.12.2016 | Online Support         | Upgrade to TIA Portal V14
     // 02.00.00 | 01.09.2017 | Online Support         | Upgrade to TIA Portal V14 SP1
     //                                                | Implementation of Programming styleguide
     //                                                | Added support for IO-Link V1.1 readers
     // 02.01.00 | 01.12.2017 | Online Support         | Bug fixes and performance improvements
     // 02.02.00 | 01.03.2020 | Online Support         | Upgrade to TIA Portal V16
     // 02.03.00 | 22.09.2020 | Online Support         | Integrated FB into LIOLink library
     //                                                | Renamed FB to LIOLink_RF200_WriteTag
     //                                                | Combined FBs for IO-Link V1.0 and V1.1
     //                                                | Minor bug fixes
     //===============================================================================
   END_REGION

   IF #version = #IOL_V11 THEN                               //determine IO-Link reader version (1.0/1.1) to set offsets
       #statIOsize := #LEN_DATA_V11;
       #statIOsizeNetto := #LEN_DATA_V11 - 4;
   ELSE
       #statIOsize := #LEN_DATA_V10;
       #statIOsizeNetto := #LEN_DATA_V10 - 4;
   END_IF;

   #statAddrOffset := #portAddr;                           //start adress of port
   #InstGetIoPart(ID     := #hwID,                              //read data from process image
                  OFFSET := #statAddrOffset,
                  LEN    := #statIOsize,
                  STATUS => #statIoPartStatus,
                  ERROR  => #statIoPartError,
                  INPUTS := #statRecDat);

   #statStatusByte := #statRecDat[0];             //Status Byte
   #statPresenceBit := #statStatusBits[5];                       //Presence bit. Transponder on field
   #presence := #statPresenceBit;

   IF NOT #execute THEN
       #statDone := false;
       #statBusy := false;
       #done := false;
       #busy := false;
       #error := false;
       #status := 0;
   ELSE
       #done := #statDone;
       #busy := #statBusy;
   END_IF;

   #statDiffToIOsizeNetto := WORD_TO_INT(#length) MOD #statIOsizeNetto;

   IF #execute AND #execute <> #statExecuteReq THEN        //Positive edge for d#reading of data
       IF NOT #statBusy THEN
           #statAddr := #addrTag;                                 //Transpoder Adress
           #statAddrTag := WORD_TO_INT(#statAddr);
           #statLength := #length;                             //Length of read Data
           #statNState := #statWriteState;
           #statBusy := TRUE;
           #statDone := FALSE;                                   //reset all the output parameters                                   
           #error := FALSE;
           #status := 0;
           #statWriteOffset := 0;
           #statBytemove := 0;
           //next step >> send write command
       ELSE
           #tempStatus_W[1] := 16#8102;                          //block is still active
           #tempStatus_W[0] := 16#0001;                          //Error identifier for block errors
           #status := #tempStatus;
           #statNState := #statErrorState;
       END_IF;
       IF #length < #statIOsizeNetto THEN
           #tempStatus_W[1] := 16#8104;                              //length too short
           #tempStatus_W[0] := 16#0001;                              //identifier rfid errors
           #status := #tempStatus;
           #statNState := #statErrorState;
       END_IF;
   END_IF;
   #statExecuteReq := #execute;

   IF NOT #presence AND #presence <> #statPresenceFf THEN   //the tag has left the antenna  field
       IF NOT #statDone THEN
           #statTimerIn := true;                              //wait 5 sec
           #statTimerR := false;
       END_IF;
   END_IF;
   #statPresenceFf := #presence;
   IF #presence THEN
       #statTimerR := true;
       #statTimerIn := false;
   END_IF;
   //-----------------------------------------------------------------------------------------------------//
   //------------------------------------------start of state machine------------------------------------//
   //-----------------------------------------------------------------------------------------------------//
   CASE #statNState OF
       0://IDLE
           #statWriteOffset := 0;                                             //offset of puffer must be reseted
           #statBusy := false;
           #statTimerIn := false;

           //-------------------------------------------------Write state-----------------------------------------//
           //---------------------------------------------send write command--------------------------------------//
           //-----------------------------------------------------------------------------------------------------//

       2://Write_state

           IF #statLength > 0 THEN
               #statDat[0] := 16#1;                      //Set write command
               #statDat[2] := #statAddrWrite[0];             //Adr-H
               #statDat[3] := #statAddrWrite[1];             //Adr-L
               VariantGet(SRC := #identData,
                          DST => #statWriteData);

               #statReturnMoveBlkVar := MOVE_BLK_VARIANT(SRC := #statWriteData,
                                                         COUNT := #statIOsizeNetto,
                                                         SRC_INDEX := #statWriteOffset - #statBytemove,
                                                         DEST_INDEX := 4,
                                                         DEST => #statDat);
               //Just #statIOsizeNetto Bytes are reserved for every transfer
           END_IF;
           IF NOT #statIoPartError THEN
               #statNState := #statTelegramState;                           //Telegram: Edit the read data
           END_IF;

           //-----------------------------------------------Telegram state----------------------------------------//
           //-----------------------------------------------------------------------------------------------------//
           //-----------------------------------------------------------------------------------------------------//  

       1://Telegram_state

           IF #statLength > 0 THEN                                  //Only when length of data>0 can continue  
               IF #statStatusBits[6] THEN                            //IF RFID error has occured
                   #tempStatus_W[1] := #statRecDat[1];
                   #tempStatus_W[0] := 16#0011;                          //Error identifier for RFID errors
                   #status := #tempStatus;
                   #statNState := #statErrorState;
               END_IF;

               //-------------------------- write command is ready------------------------------------------------//

               IF #statStatusBits[7] AND #statStatusBits[0] THEN
                   IF #statRecDat[2] = #statAddrWrite[0] AND #statRecDat[3] = #statAddrWrite[1] THEN //received ADR must be ==sent ADR

                       IF NOT #statIoPartError THEN
                           IF #statStatusBits[7] AND NOT #statStatusBits[6] THEN
                               #statLength := #statLength - #statIOsizeNetto;
                               IF #statDiffToIOsizeNetto <> 0 AND #statLength < #statIOsizeNetto THEN
                                   #statBytemove := #statIOsizeNetto - #statDiffToIOsizeNetto;
                               END_IF;
                               //if len is not dividable with #statIOsizeNetto the adr offset has to be changed that the last (length < #statIOsizeNetto) command is done right
                               #statWriteOffset := #statWriteOffset + #statIOsizeNetto;                                   //offset must be changed
                               #statAddr := INT_TO_WORD(WORD_TO_INT(#statAddr) + #statIOsizeNetto) - INT_TO_WORD(#statBytemove);     //Change the ADR on Transponder(#statIOsizeNetto Bytes)       
                               #statNState := #statWriteState;                      //Start a new write command
                           ELSE
                               #statNState := #statIdleState;
                           END_IF;
                       ELSE
                           #tempStatus_W[1] := DWORD_TO_WORD(#statIoPartStatus);                 //Error has to BLKMOV occured
                           #tempStatus_W[0] := 16#0001;                           //functions-Error identifier
                           #status := #tempStatus;
                           #statNState := #statErrorState;
                       END_IF;
                   END_IF;
               END_IF;

               #InstSetIoPart(ID      := #hwID,
                              OFFSET  := #statAddrOffset,
                              LEN     := #statIOsize,
                              STATUS  => #statIoPartStatus,
                              ERROR   => #statIoPartError,
                              OUTPUTS := #statDat);

               IF #statIoPartError THEN
                   #tempStatus_W[1] := DWORD_TO_WORD(#statIoPartStatus);   //Error has to BLKMOV occured
                   #tempStatus_W[0] := 16#0001;                            //functions-Error identifier
                   #status := #tempStatus;
                   #statNState := #statErrorState;
               END_IF;

           ELSE
               #statNState := #statIdleState;
               #statBusy := false;
               #statDone := TRUE;

               //Reset write command
               #statDat[0] := 16#0;

               #InstSetIoPart(ID      := #hwID,
                              OFFSET  := #statAddrOffset,
                              LEN     := #statIOsize,
                              STATUS  => #statIoPartStatus,
                              ERROR   => #statIoPartError,
                              OUTPUTS := #statDat);
           END_IF;

           //------------------------------------------------------------------------------------------------------------//
           //-------------------------------------------------Error state------------------------------------------------//
           //---------------------------------------------error has occured----------------------------------------------//

       3://Error_State
           #tempError := TRUE;
           #statBusy := false;
           #error := #tempError;
           #statDone := false;
           #statTimerIn := false;
           #statTimerR := true;
           #statNState := #statIdleState;

           //Reset write command
           #statDat[0] := 16#0;

           #InstSetIoPart(ID      := #hwID,
                          OFFSET  := #statAddrOffset,
                          LEN     := #statIOsize,
                          STATUS  => #statIoPartStatus,
                          ERROR   => #statIoPartError,
                          OUTPUTS := #statDat);
   END_CASE;


   //------------------------------------------------------------------------------------------------------------//
   //-------------------------------------------------Timer------------------------------------------------------//
   //------------------------------------------------------------------------------------------------------------//

   #instTonR(IN := #statTimerIn,               //this timer will start, if the tag has left the antenna field
             R  := #statTimerR,
             PT := #statTimerPt);
   IF #instTonR.Q THEN                      //error has occured. No tag on field during the 5 sec.
       #tempStatus_W[1] := 16#8101;                              //tag has left the field
       #tempStatus_W[0] := 16#0001;                              //identifier rfid errors
       #status := #tempStatus;
       #statNState := #statErrorState;
   END_IF;
END_FUNCTION_BLOCK

(* ===== HMI "HMI_RT_1" =====
connection "HMI_Connection_1": ETHERNET, S7_1500_OMS

HMI tags "Default tag table"
   "DB_MES_Comms_station_state" : Int = PLC DB_MES_Comms.station_state, 100 ms
   "DB_MES_Comms_good_count" : Int = PLC DB_MES_Comms.good_count, 100 ms
   "DB_MES_Comms_total_count" : Int = PLC DB_MES_Comms.total_count, 100 ms
   "start" : Bool = PLC start AT %I1.0, 100 ms
   "stop" : Bool = PLC stop AT %I1.1, 1 s
   "reset" : Bool = PLC reset AT %I1.3, 1 s
   "conv_start" : Bool = PLC conv_start AT %I1.6, 1 s
   "conv_centre" : Bool = PLC conv_centre AT %I1.4, 1 s
   "conv_end" : Bool = PLC conv_end AT %I1.7, 1 s
   "F1_F2" : Bool = PLC F1_F2 AT %I1.2, 1 s

text list "Station_State_Display": 1 'ACTIVE'; 2 'DONE'; 0 'IDLE'

screen "Screen_1" 800x480
   TextField "Text field_1" at 357,8 size 122x23; Text 'LabelProMax'
   TextField "Text field_2" at 62,73 size 16x23; Text 'Text'
   TextField "Text field_6" at 51,162 size 152x23; Text 'STATION STATE'
   Button "Button_1" at 19,59 size 166x60; TextOff 'START'
      Appearance <- "start"
   Button "Button_2" at 203,59 size 166x60; TextOff 'STOP'
      Appearance <- "stop"
   Button "Button_3" at 407,59 size 166x60; TextOff 'RESET'
      Appearance <- "reset"
   Switch "Switch_2" at 619,40 size 120x88; CaptionText 'MODE'; TextOff 'F2'; TextOn 'F1'
      ObjectEnable <- "F1_F2"
   TextField "Text field_3" at 324,162 size 126x23; Text 'GOOD COUNT'
   IOField "I/O field_2" at 314,210 size 136x48; FormatPattern s99999
      ProcessValue <- "DB_MES_Comms_good_count"
   IOField "I/O field_3" at 586,212 size 136x48; FormatPattern s99999
      ProcessValue <- "DB_MES_Comms_total_count"
   TextField "Text field_4" at 596,162 size 134x23; Text 'TOTAL COUNT'
   SymbolicIOField "Symbolic I/O field_1" at 34,218 size 170x32; TextOff '0'; TextOn '1'; TextList "Station_State_Display"
      ProcessValue <- "DB_MES_Comms_station_state"
   Circle "Circle_3" at 49,408 size 29x29
      Appearance <- "conv_start"
   Circle "Circle_4" at 369,408 size 29x29
      Appearance <- "conv_centre"
   Circle "Circle_5" at 689,408 size 29x29
      Appearance <- "conv_end"
   TextField "Text field_5" at 41,437 size 51x23; Text 'Start'
   TextField "Text field_8" at 340,437 size 88x23; Text 'Labelling'
   TextField "Text field_9" at 686,437 size 38x23; Text 'End'
   TextField "Text field_10" at 42,275 size 228x23; Text 'Conveyor Belt Visualizer'
   Group "Group" at 62,328 size 96x48
   Group "Group_1" at 340,328 size 96x48
   Group "Group_2" at 619,328 size 96x48
   Rectangle "Rectangle_7" at 62,328 size 96x48
      Visibility <- "conv_start"
   Rectangle "Rectangle_8" at 72,334 size 74x36
      Visibility <- "conv_start"
   Rectangle "Rectangle_9" at 340,328 size 96x48
      Visibility <- "conv_centre"
   Rectangle "Rectangle_10" at 350,334 size 74x36
      Visibility <- "conv_centre"
   Rectangle "Rectangle_11" at 619,328 size 96x48
      Visibility <- "conv_end"
   Rectangle "Rectangle_12" at 629,334 size 74x36
      Visibility <- "conv_end"
*)